screen "Point_1" 800x480, template "Main"
   TextField "Text field_1" at 0,2 size 547x23; Text 'Таблица настройки зависимостей дозы от мутность для линии 1'
   TextField "Text field_12" at 566,23 size 71x23; Text 'Запрос:'
   IOField "I/O field_4" at 653,22 size 66x25; FormatPattern 999.99
      ProcessValue <- "Ponts_1_DB_REQ"
   TextField "Text field_4" at 566,46 size 84x23; Text 'Команда:'
   IOField "I/O field_2" at 653,45 size 66x25; FormatPattern 999.99
      ProcessValue <- "Ponts_1_DB_Value"
   TextField "Text field_40" at 566,69 size 84x23; Text 'Датчик:'
   IOField "I/O field_24" at 653,68 size 66x25; FormatPattern 999.99
      ProcessValue <- "AIx_DB_Trans_1_Result"
   Rectangle "Rectangle_1" at 142,113 size 111x147
      Appearance <- "Ponts_1_DB_Now{1}"
   TextField "Text field_3" at 164,141 size 67x20; Text 'мутность'
   TextField "Text field_5" at 179,196 size 37x20; Text 'доза'
   TextField "Text field_11" at 142,115 size 95x25; Text 'Точка 1'
   Button "Button_1" at 223,113 size 30x30; TextOff 'Text'; Authorization "Operator"; PictureList "on_off_1"
      on Click: InvertBit("Ponts_1_DB_PLF_1_Use")
      ProcessValue <- "Ponts_1_DB_PLF_1_Use"
   IOField "I/O field_16" at 157,160 size 82x40; Authorization "Operator"; FormatPattern 999.99
      ProcessValue <- "Ponts_1_DB_PLF_1_High"
   IOField "I/O field_17" at 157,216 size 82x40; Authorization "Operator"; FormatPattern 999.99
      ProcessValue <- "Ponts_1_DB_PLF_1_Point_B"
   TextField "Text field_9" at 2,35 size 164x23; Text 'Минимальная доза'
   TextField "Text field_10" at 2,64 size 172x23; Text 'Максимальная доза'
   IOField "I/O field_1" at 181,33 size 70x30; Authorization "Operator"; FormatPattern 999.99
      ProcessValue <- "Ponts_1_DB_Min"
   IOField "I/O field_30" at 181,64 size 70x30; Authorization "Operator"; FormatPattern 999.99
      ProcessValue <- "Ponts_1_DB_Max"
   Rectangle "Rectangle_2" at 21,113 size 111x147
      Appearance <- "Ponts_1_DB_Now{0}"
   TextField "Text field_2" at 43,141 size 67x20; Text 'мутность'
   TextField "Text field_6" at 58,196 size 37x20; Text 'доза'
   TextField "Text field_7" at 21,115 size 95x25; Text 'Точка 0'
   Button "Button_2" at 102,113 size 30x30; TextOff 'Text'; Authorization "Operator"; PictureList "on_off_1"
      on Click: InvertBit("Ponts_1_DB_PLF_0_Use")
      ProcessValue <- "Ponts_1_DB_PLF_0_Use"
   IOField "I/O field_3" at 36,160 size 82x40; Authorization "Operator"; FormatPattern 999.99
      ProcessValue <- "Ponts_1_DB_PLF_0_High"
   IOField "I/O field_5" at 36,216 size 82x40; Authorization "Operator"; FormatPattern 999.99
      ProcessValue <- "Ponts_1_DB_PLF_0_Point_B"
   Rectangle "Rectangle_3" at 264,114 size 111x147
      Appearance <- "Ponts_1_DB_Now{2}"
   TextField "Text field_8" at 286,142 size 67x20; Text 'мутность'
   TextField "Text field_13" at 301,197 size 37x20; Text 'доза'
   TextField "Text field_14" at 264,116 size 95x25; Text 'Точка 2'
   Button "Button_3" at 345,114 size 30x30; TextOff 'Text'; Authorization "Operator"; PictureList "on_off_1"
      on Click: InvertBit("Ponts_1_DB_PLF_2_Use")
      ProcessValue <- "Ponts_1_DB_PLF_2_Use"
   IOField "I/O field_6" at 279,161 size 82x40; Authorization "Operator"; FormatPattern 999.99
      ProcessValue <- "Ponts_1_DB_PLF_2_High"
   IOField "I/O field_7" at 279,217 size 82x40; Authorization "Operator"; FormatPattern 999.99
      ProcessValue <- "Ponts_1_DB_PLF_2_Point_B"
   Rectangle "Rectangle_4" at 386,115 size 111x147
      Appearance <- "Ponts_1_DB_Now{3}"
   TextField "Text field_15" at 408,143 size 67x20; Text 'мутность'
   TextField "Text field_16" at 423,198 size 37x20; Text 'доза'
   TextField "Text field_17" at 386,117 size 95x25; Text 'Точка 3'
   Button "Button_4" at 467,115 size 30x30; TextOff 'Text'; Authorization "Operator"; PictureList "on_off_1"
      on Click: InvertBit("Ponts_1_DB_PLF_3_Use")
      ProcessValue <- "Ponts_1_DB_PLF_3_Use"
   IOField "I/O field_8" at 401,162 size 82x40; Authorization "Operator"; FormatPattern 999.99
      ProcessValue <- "Ponts_1_DB_PLF_3_High"
   IOField "I/O field_9" at 401,218 size 82x40; Authorization "Operator"; FormatPattern 999.99
      ProcessValue <- "Ponts_1_DB_PLF_3_Point_B"
   Rectangle "Rectangle_5" at 142,287 size 111x147
      Appearance <- "Ponts_1_DB_Now{5}"
   TextField "Text field_18" at 164,315 size 67x20; Text 'мутность'
   TextField "Text field_19" at 179,370 size 37x20; Text 'доза'
   TextField "Text field_20" at 142,289 size 95x25; Text 'Точка 5'
   Button "Button_5" at 223,287 size 30x30; TextOff 'Text'; Authorization "Operator"; PictureList "on_off_1"
      on Click: InvertBit("Ponts_1_DB_PLF_5_Use")
      ProcessValue <- "Ponts_1_DB_PLF_5_Use"
   IOField "I/O field_10" at 157,334 size 82x40; Authorization "Operator"; FormatPattern 999.99
      ProcessValue <- "Ponts_1_DB_PLF_5_High"
   IOField "I/O field_11" at 157,390 size 82x40; Authorization "Operator"; FormatPattern 999.99
      ProcessValue <- "Ponts_1_DB_PLF_5_Point_B"
   Rectangle "Rectangle_6" at 21,287 size 111x147
      Appearance <- "Ponts_1_DB_Now{4}"
   TextField "Text field_21" at 43,315 size 67x20; Text 'мутность'
   TextField "Text field_22" at 58,370 size 37x20; Text 'доза'
   TextField "Text field_23" at 21,289 size 95x25; Text 'Точка 4'
   Button "Button_6" at 102,287 size 30x30; TextOff 'Text'; Authorization "Operator"; PictureList "on_off_1"
      on Click: InvertBit("Ponts_1_DB_PLF_4_Use")
      ProcessValue <- "Ponts_1_DB_PLF_4_Use"
   IOField "I/O field_12" at 36,334 size 82x40; Authorization "Operator"; FormatPattern 999.99
      ProcessValue <- "Ponts_1_DB_PLF_4_High"
   IOField "I/O field_13" at 36,390 size 82x40; Authorization "Operator"; FormatPattern 999.99
      ProcessValue <- "Ponts_1_DB_PLF_4_Point_B"
   Rectangle "Rectangle_7" at 264,288 size 111x147
      Appearance <- "Ponts_1_DB_Now{6}"
   TextField "Text field_24" at 286,316 size 67x20; Text 'мутность'
   TextField "Text field_25" at 301,371 size 37x20; Text 'доза'
   TextField "Text field_26" at 264,290 size 95x25; Text 'Точка 6'
   Button "Button_7" at 345,288 size 30x30; TextOff 'Text'; Authorization "Operator"; PictureList "on_off_1"
      on Click: InvertBit("Ponts_1_DB_PLF_6_Use")
      ProcessValue <- "Ponts_1_DB_PLF_6_Use"
   IOField "I/O field_14" at 279,335 size 82x40; Authorization "Operator"; FormatPattern 999.99
      ProcessValue <- "Ponts_1_DB_PLF_6_High"
   IOField "I/O field_15" at 279,391 size 82x40; Authorization "Operator"; FormatPattern 999.99
      ProcessValue <- "Ponts_1_DB_PLF_6_Point_B"
   Rectangle "Rectangle_8" at 386,289 size 111x147
      Appearance <- "Ponts_1_DB_Now{7}"
   TextField "Text field_27" at 408,317 size 67x20; Text 'мутность'
   TextField "Text field_28" at 423,372 size 37x20; Text 'доза'
   TextField "Text field_29" at 386,291 size 95x25; Text 'Точка 7'
   Button "Button_8" at 467,289 size 30x30; TextOff 'Text'; Authorization "Operator"; PictureList "on_off_1"
      on Click: InvertBit("Ponts_1_DB_PLF_7_Use")
      ProcessValue <- "Ponts_1_DB_PLF_7_Use"
   IOField "I/O field_18" at 401,336 size 82x40; Authorization "Operator"; FormatPattern 999.99
      ProcessValue <- "Ponts_1_DB_PLF_7_High"
   IOField "I/O field_19" at 401,392 size 82x40; Authorization "Operator"; FormatPattern 999.99
      ProcessValue <- "Ponts_1_DB_PLF_7_Point_B"

screen "Point_2" 800x480, template "Main"
   TextField "Text field_1" at 0,2 size 547x23; Text 'Таблица настройки зависимостей дозы от мутность для линии 2'
   TextField "Text field_12" at 566,23 size 71x23; Text 'Запрос:'
   IOField "I/O field_4" at 653,22 size 66x25; FormatPattern 999.99
      ProcessValue <- "Ponts_2_DB_REQ"
   TextField "Text field_4" at 566,46 size 84x23; Text 'Команда:'
   IOField "I/O field_2" at 653,45 size 66x25; FormatPattern 999.99
      ProcessValue <- "Ponts_2_DB_Value"
   TextField "Text field_40" at 566,69 size 84x23; Text 'Датчик:'
   IOField "I/O field_24" at 653,68 size 66x25; FormatPattern 999.99
      ProcessValue <- "AIx_DB_Trans_2_Result"
   Rectangle "Rectangle_1" at 142,113 size 111x147
      Appearance <- "Ponts_2_DB_Now{1}"
   TextField "Text field_3" at 164,141 size 67x20; Text 'мутность'
   TextField "Text field_5" at 179,196 size 37x20; Text 'доза'
   TextField "Text field_11" at 142,115 size 95x25; Text 'Точка 1'
   Button "Button_1" at 223,113 size 30x30; TextOff 'Text'; Authorization "Operator"; PictureList "on_off_1"
      on Click: InvertBit("Ponts_2_DB_PLF_1_Use")
      ProcessValue <- "Ponts_2_DB_PLF_1_Use"
   IOField "I/O field_16" at 157,160 size 82x40; Authorization "Operator"; FormatPattern 999.99
      ProcessValue <- "Ponts_2_DB_PLF_1_High"
   IOField "I/O field_17" at 157,216 size 82x40; Authorization "Operator"; FormatPattern 999.99
      ProcessValue <- "Ponts_2_DB_PLF_1_Point_B"
   TextField "Text field_9" at 2,35 size 164x23; Text 'Минимальная доза'
   TextField "Text field_10" at 2,64 size 172x23; Text 'Максимальная доза'
   IOField "I/O field_1" at 181,33 size 70x30; Authorization "Operator"; FormatPattern 999.99
      ProcessValue <- "Ponts_2_DB_Min"
   IOField "I/O field_30" at 181,64 size 70x30; Authorization "Operator"; FormatPattern 999.99
      ProcessValue <- "Ponts_2_DB_Max"
   Rectangle "Rectangle_2" at 21,113 size 111x147
      Appearance <- "Ponts_2_DB_Now{0}"
   TextField "Text field_2" at 43,141 size 67x20; Text 'мутность'
   TextField "Text field_6" at 58,196 size 37x20; Text 'доза'
   TextField "Text field_7" at 21,115 size 95x25; Text 'Точка 0'
   Button "Button_2" at 102,113 size 30x30; TextOff 'Text'; Authorization "Operator"; PictureList "on_off_1"
      on Click: InvertBit("Ponts_2_DB_PLF_0_Use")
      ProcessValue <- "Ponts_2_DB_PLF_0_Use"
   IOField "I/O field_3" at 36,160 size 82x40; Authorization "Operator"; FormatPattern 999.99
      ProcessValue <- "Ponts_2_DB_PLF_0_High"
   IOField "I/O field_5" at 36,216 size 82x40; Authorization "Operator"; FormatPattern 999.99
      ProcessValue <- "Ponts_2_DB_PLF_0_Point_B"
   Rectangle "Rectangle_3" at 264,114 size 111x147
      Appearance <- "Ponts_2_DB_Now{2}"
   TextField "Text field_8" at 286,142 size 67x20; Text 'мутность'
   TextField "Text field_13" at 301,197 size 37x20; Text 'доза'
   TextField "Text field_14" at 264,116 size 95x25; Text 'Точка 2'
   Button "Button_3" at 345,114 size 30x30; TextOff 'Text'; Authorization "Operator"; PictureList "on_off_1"
      on Click: InvertBit("Ponts_2_DB_PLF_2_Use")
      ProcessValue <- "Ponts_2_DB_PLF_2_Use"
   IOField "I/O field_6" at 279,161 size 82x40; Authorization "Operator"; FormatPattern 999.99
      ProcessValue <- "Ponts_2_DB_PLF_2_High"
   IOField "I/O field_7" at 279,217 size 82x40; Authorization "Operator"; FormatPattern 999.99
      ProcessValue <- "Ponts_2_DB_PLF_2_Point_B"
   Rectangle "Rectangle_4" at 386,115 size 111x147
      Appearance <- "Ponts_2_DB_Now{3}"
   TextField "Text field_15" at 408,143 size 67x20; Text 'мутность'
   TextField "Text field_16" at 423,198 size 37x20; Text 'доза'
   TextField "Text field_17" at 386,117 size 95x25; Text 'Точка 3'
   Button "Button_4" at 467,115 size 30x30; TextOff 'Text'; Authorization "Operator"; PictureList "on_off_1"
      on Click: InvertBit("Ponts_2_DB_PLF_3_Use")
      ProcessValue <- "Ponts_2_DB_PLF_3_Use"
   IOField "I/O field_8" at 401,162 size 82x40; Authorization "Operator"; FormatPattern 999.99
      ProcessValue <- "Ponts_2_DB_PLF_3_High"
   IOField "I/O field_9" at 401,218 size 82x40; Authorization "Operator"; FormatPattern 999.99
      ProcessValue <- "Ponts_2_DB_PLF_3_Point_B"
   Rectangle "Rectangle_5" at 142,287 size 111x147
      Appearance <- "Ponts_2_DB_Now{5}"
   TextField "Text field_18" at 164,315 size 67x20; Text 'мутность'
   TextField "Text field_19" at 179,370 size 37x20; Text 'доза'
   TextField "Text field_20" at 142,289 size 95x25; Text 'Точка 5'
   Button "Button_5" at 223,287 size 30x30; TextOff 'Text'; Authorization "Operator"; PictureList "on_off_1"
      on Click: InvertBit("Ponts_2_DB_PLF_5_Use")
      ProcessValue <- "Ponts_2_DB_PLF_5_Use"
   IOField "I/O field_10" at 157,334 size 82x40; Authorization "Operator"; FormatPattern 999.99
      ProcessValue <- "Ponts_2_DB_PLF_5_High"
   IOField "I/O field_11" at 157,390 size 82x40; Authorization "Operator"; FormatPattern 999.99
      ProcessValue <- "Ponts_2_DB_PLF_5_Point_B"
   Rectangle "Rectangle_6" at 21,287 size 111x147
      Appearance <- "Ponts_2_DB_Now{4}"
   TextField "Text field_21" at 43,315 size 67x20; Text 'мутность'
   TextField "Text field_22" at 58,370 size 37x20; Text 'доза'
   TextField "Text field_23" at 21,289 size 95x25; Text 'Точка 4'
   Button "Button_6" at 102,287 size 30x30; TextOff 'Text'; Authorization "Operator"; PictureList "on_off_1"
      on Click: InvertBit("Ponts_2_DB_PLF_4_Use")
      ProcessValue <- "Ponts_2_DB_PLF_4_Use"
   IOField "I/O field_12" at 36,334 size 82x40; Authorization "Operator"; FormatPattern 999.99
      ProcessValue <- "Ponts_2_DB_PLF_4_High"
   IOField "I/O field_13" at 36,390 size 82x40; Authorization "Operator"; FormatPattern 999.99
      ProcessValue <- "Ponts_2_DB_PLF_4_Point_B"
   Rectangle "Rectangle_7" at 264,288 size 111x147
      Appearance <- "Ponts_2_DB_Now{6}"
   TextField "Text field_24" at 286,316 size 67x20; Text 'мутность'
   TextField "Text field_25" at 301,371 size 37x20; Text 'доза'
   TextField "Text field_26" at 264,290 size 95x25; Text 'Точка 6'
   Button "Button_7" at 345,288 size 30x30; TextOff 'Text'; Authorization "Operator"; PictureList "on_off_1"
      on Click: InvertBit("Ponts_2_DB_PLF_6_Use")
      ProcessValue <- "Ponts_2_DB_PLF_6_Use"
   IOField "I/O field_14" at 279,335 size 82x40; Authorization "Operator"; FormatPattern 999.99
      ProcessValue <- "Ponts_2_DB_PLF_6_High"
   IOField "I/O field_15" at 279,391 size 82x40; Authorization "Operator"; FormatPattern 999.99
      ProcessValue <- "Ponts_2_DB_PLF_6_Point_B"
   Rectangle "Rectangle_8" at 386,289 size 111x147
      Appearance <- "Ponts_2_DB_Now{7}"
   TextField "Text field_27" at 408,317 size 67x20; Text 'мутность'
   TextField "Text field_28" at 423,372 size 37x20; Text 'доза'
   TextField "Text field_29" at 386,291 size 95x25; Text 'Точка 7'
   Button "Button_8" at 467,289 size 30x30; TextOff 'Text'; Authorization "Operator"; PictureList "on_off_1"
      on Click: InvertBit("Ponts_2_DB_PLF_7_Use")
      ProcessValue <- "Ponts_2_DB_PLF_7_Use"
   IOField "I/O field_18" at 401,336 size 82x40; Authorization "Operator"; FormatPattern 999.99
      ProcessValue <- "Ponts_2_DB_PLF_7_High"
   IOField "I/O field_19" at 401,392 size 82x40; Authorization "Operator"; FormatPattern 999.99
      ProcessValue <- "Ponts_2_DB_PLF_7_Point_B"

screen "Mass_1" 800x480, template "Main"
   TextField "Text field_1" at 220,5 size 368x47; Text 'Статистика весов 1'
   Button "HmiScreenItemData_1" at 10,425 size 159x47; TextOn 'Система'; TextOff 'Прошлый месяц'; PictureOn "Navigates to System screens for KTP700 Basic+ PN 14.0.1.0"; PictureOff "Navigates to System screens for KTP700 Basic+ PN 14.0.1.0"
      on Release: ActivateScreen("Last_1", 0)
   Button "HmiScreenItemData_4" at 565,425 size 159x47; TextOn 'О нас'; TextOff 'Текущий месяц'; PictureOn "Navigates to System screens for KTP700 Basic+ PN 14.0.1.0"; PictureOff "Navigates to System screens for KTP700 Basic+ PN 14.0.1.0"
   IOField "I/O field_1" at 365,434 size 98x30; FormatPattern 99999.99
      ProcessValue <- "Statistics_DB_Today_1"
      Appearance <- "DIx_DB_Mass_1_Signal"
   TextField "Text field_17" at 257,435 size 93x27; Text 'Сегодня:'
   TextField "Text field_2" at 10,5 size 75x23; Text 'Сегодня'
   TextField "Text field_3" at 126,5 size 45x23; Text 'день'
   IOField "I/O field_2" at 88,3 size 37x30; FormatPattern 99
      ProcessValue <- "Statistics_DB_Today_Int"
      Appearance <- "DIx_DB_Mass_1_Signal"
   TextField "Text field_4" at 12,61 size 61x23; Text 'День 1'
   TextField "Text field_5" at 12,97 size 61x23; Text 'День 2'
   TextField "Text field_6" at 12,134 size 61x23; Text 'День 3'
   TextField "Text field_7" at 12,170 size 61x23; Text 'День 4'
   TextField "Text field_8" at 12,207 size 61x23; Text 'День 5'
   TextField "Text field_9" at 12,243 size 61x23; Text 'День 6'
   TextField "Text field_10" at 12,280 size 61x23; Text 'День 7'
   TextField "Text field_11" at 12,316 size 61x23; Text 'День 8'
   TextField "Text field_12" at 12,353 size 61x23; Text 'День 9'
   TextField "Text field_13" at 12,390 size 71x23; Text 'День 10'
   IOField "I/O field_8" at 90,59 size 80x27; Authorization "Operator"; FormatPattern 999999.9
      ProcessValue <- "Statistics_DB_Month_1{1}"
   IOField "I/O field_3" at 90,95 size 80x27; Authorization "Operator"; FormatPattern 999999.9
      ProcessValue <- "Statistics_DB_Month_1{2}"
   IOField "I/O field_4" at 90,132 size 80x27; Authorization "Operator"; FormatPattern 999999.9
      ProcessValue <- "Statistics_DB_Month_1{3}"
   IOField "I/O field_5" at 90,168 size 80x27; Authorization "Operator"; FormatPattern 999999.9
      ProcessValue <- "Statistics_DB_Month_1{4}"
   IOField "I/O field_6" at 90,205 size 80x27; Authorization "Operator"; FormatPattern 999999.9
      ProcessValue <- "Statistics_DB_Month_1{5}"
   IOField "I/O field_7" at 90,241 size 80x27; Authorization "Operator"; FormatPattern 999999.9
      ProcessValue <- "Statistics_DB_Month_1{6}"
   IOField "I/O field_9" at 90,278 size 80x27; Authorization "Operator"; FormatPattern 999999.9
      ProcessValue <- "Statistics_DB_Month_1{7}"
   IOField "I/O field_10" at 90,314 size 80x27; Authorization "Operator"; FormatPattern 999999.9
      ProcessValue <- "Statistics_DB_Month_1{8}"
   IOField "I/O field_11" at 90,351 size 80x27; Authorization "Operator"; FormatPattern 999999.9
      ProcessValue <- "Statistics_DB_Month_1{9}"
   IOField "I/O field_12" at 90,388 size 80x27; Authorization "Operator"; FormatPattern 999999.9
      ProcessValue <- "Statistics_DB_Month_1{10}"
   IOField "I/O field_13" at 565,316 size 159x30; FormatPattern 99999.9
      ProcessValue <- "Statistics_DB_Summ_1"
      Appearance <- "DIx_DB_Mass_1_Signal"
   TextField "Text field_14" at 595,284 size 100x27; Text 'За месяц:'
   TextField "Text field_15" at 611,359 size 67x27; Text 'Всего:'
   IOField "I/O field_14" at 565,387 size 159x30; FormatPattern 9999999.9
      ProcessValue <- "Statistics_DB_All_1"
      Appearance <- "DIx_DB_Mass_1_Signal"
   TextField "Text field_16" at 202,62 size 71x23; Text 'День 11'
   TextField "Text field_18" at 202,98 size 71x23; Text 'День 12'
   TextField "Text field_19" at 202,135 size 71x23; Text 'День 13'
   TextField "Text field_20" at 202,171 size 71x23; Text 'День 14'
   TextField "Text field_21" at 202,208 size 71x23; Text 'День 15'
   TextField "Text field_22" at 202,244 size 71x23; Text 'День 16'
   TextField "Text field_23" at 202,281 size 71x23; Text 'День 17'
   TextField "Text field_24" at 202,317 size 71x23; Text 'День 18'
   TextField "Text field_25" at 202,354 size 71x23; Text 'День 19'
   TextField "Text field_26" at 202,391 size 71x23; Text 'День 20'
   IOField "I/O field_15" at 280,60 size 80x27; Authorization "Operator"; FormatPattern 999999.9
      ProcessValue <- "Statistics_DB_Month_1{11}"
   IOField "I/O field_16" at 280,96 size 80x27; Authorization "Operator"; FormatPattern 999999.9
      ProcessValue <- "Statistics_DB_Month_1{12}"
   IOField "I/O field_17" at 280,133 size 80x27; Authorization "Operator"; FormatPattern 999999.9
      ProcessValue <- "Statistics_DB_Month_1{13}"
   IOField "I/O field_18" at 280,169 size 80x27; Authorization "Operator"; FormatPattern 999999.9
      ProcessValue <- "Statistics_DB_Month_1{14}"
   IOField "I/O field_19" at 280,206 size 80x27; Authorization "Operator"; FormatPattern 999999.9
      ProcessValue <- "Statistics_DB_Month_1{15}"
   IOField "I/O field_20" at 280,242 size 80x27; Authorization "Operator"; FormatPattern 999999.9
      ProcessValue <- "Statistics_DB_Month_1{16}"
   IOField "I/O field_21" at 280,279 size 80x27; Authorization "Operator"; FormatPattern 999999.9
      ProcessValue <- "Statistics_DB_Month_1{17}"
   IOField "I/O field_22" at 280,315 size 80x27; Authorization "Operator"; FormatPattern 999999.9
      ProcessValue <- "Statistics_DB_Month_1{18}"
   IOField "I/O field_23" at 280,352 size 80x27; Authorization "Operator"; FormatPattern 999999.9
      ProcessValue <- "Statistics_DB_Month_1{19}"
   IOField "I/O field_24" at 280,389 size 80x27; Authorization "Operator"; FormatPattern 999999.9
      ProcessValue <- "Statistics_DB_Month_1{20}"
   TextField "Text field_27" at 392,63 size 71x23; Text 'День 21'
   TextField "Text field_28" at 392,99 size 71x23; Text 'День 22'
   TextField "Text field_29" at 392,136 size 71x23; Text 'День 23'
   TextField "Text field_30" at 392,172 size 71x23; Text 'День 24'
   TextField "Text field_31" at 392,209 size 71x23; Text 'День 25'
   TextField "Text field_32" at 392,245 size 71x23; Text 'День 26'
   TextField "Text field_33" at 392,282 size 71x23; Text 'День 27'
   TextField "Text field_34" at 392,318 size 71x23; Text 'День 28'
   TextField "Text field_35" at 392,355 size 71x23; Text 'День 29'
   TextField "Text field_36" at 392,392 size 71x23; Text 'День 30'
   IOField "I/O field_25" at 470,61 size 80x27; Authorization "Operator"; FormatPattern 999999.9
      ProcessValue <- "Statistics_DB_Month_1{21}"
   IOField "I/O field_26" at 470,97 size 80x27; Authorization "Operator"; FormatPattern 999999.9
      ProcessValue <- "Statistics_DB_Month_1{22}"
   IOField "I/O field_27" at 470,134 size 80x27; Authorization "Operator"; FormatPattern 999999.9
      ProcessValue <- "Statistics_DB_Month_1{23}"
   IOField "I/O field_28" at 470,170 size 80x27; Authorization "Operator"; FormatPattern 999999.9
      ProcessValue <- "Statistics_DB_Month_1{24}"
   IOField "I/O field_29" at 470,207 size 80x27; Authorization "Operator"; FormatPattern 999999.9
      ProcessValue <- "Statistics_DB_Month_1{25}"
   IOField "I/O field_30" at 470,243 size 80x27; Authorization "Operator"; FormatPattern 999999.9
      ProcessValue <- "Statistics_DB_Month_1{26}"
   IOField "I/O field_31" at 470,280 size 80x27; Authorization "Operator"; FormatPattern 999999.9
      ProcessValue <- "Statistics_DB_Month_1{27}"
   IOField "I/O field_32" at 470,316 size 80x27; Authorization "Operator"; FormatPattern 999999.9
      ProcessValue <- "Statistics_DB_Month_1{28}"
   IOField "I/O field_33" at 470,353 size 80x27; Authorization "Operator"; FormatPattern 999999.9
      ProcessValue <- "Statistics_DB_Month_1{29}"
   IOField "I/O field_34" at 470,390 size 80x27; Authorization "Operator"; FormatPattern 999999.9
      ProcessValue <- "Statistics_DB_Month_1{30}"
   TextField "Text field_37" at 563,64 size 71x23; Text 'День 31'
   IOField "I/O field_35" at 644,62 size 80x27; Authorization "Operator"; FormatPattern 999999.9
      ProcessValue <- "Statistics_DB_Month_1{31}"

screen "Mass_2" 800x480, template "Main"
   TextField "Text field_1" at 220,5 size 368x47; Text 'Статистика весов 2'
   Button "HmiScreenItemData_1" at 10,425 size 159x47; TextOn 'Система'; TextOff 'Прошлый месяц'; PictureOn "Navigates to System screens for KTP700 Basic+ PN 14.0.1.0"; PictureOff "Navigates to System screens for KTP700 Basic+ PN 14.0.1.0"
      on Release: ActivateScreen("Last_2", 0)
   Button "HmiScreenItemData_4" at 565,425 size 159x47; TextOn 'О нас'; TextOff 'Текущий месяц'; PictureOn "Navigates to System screens for KTP700 Basic+ PN 14.0.1.0"; PictureOff "Navigates to System screens for KTP700 Basic+ PN 14.0.1.0"
   IOField "I/O field_1" at 365,434 size 98x30; FormatPattern 99999.99
      ProcessValue <- "Statistics_DB_Today_2"
      Appearance <- "DIx_DB_Mass_2_Signal"
   TextField "Text field_17" at 257,435 size 93x27; Text 'Сегодня:'
   TextField "Text field_3" at 10,5 size 75x23; Text 'Сегодня'
   TextField "Text field_4" at 126,5 size 45x23; Text 'день'
   IOField "I/O field_2" at 88,3 size 37x30; FormatPattern 99
      ProcessValue <- "Statistics_DB_Today_Int"
      Appearance <- "DIx_DB_Mass_1_Signal"
   TextField "Text field_5" at 12,61 size 61x23; Text 'День 1'
   TextField "Text field_6" at 12,97 size 61x23; Text 'День 2'
   TextField "Text field_7" at 12,134 size 61x23; Text 'День 3'
   TextField "Text field_8" at 12,170 size 61x23; Text 'День 4'
   TextField "Text field_9" at 12,207 size 61x23; Text 'День 5'
   TextField "Text field_10" at 12,243 size 61x23; Text 'День 6'
   TextField "Text field_11" at 12,280 size 61x23; Text 'День 7'
   TextField "Text field_12" at 12,316 size 61x23; Text 'День 8'
   TextField "Text field_13" at 12,353 size 61x23; Text 'День 9'
   TextField "Text field_14" at 12,390 size 71x23; Text 'День 10'
   IOField "I/O field_8" at 90,59 size 80x27; Authorization "Operator"; FormatPattern 999999.9
      ProcessValue <- "Statistics_DB_Month_2{1}"
   IOField "I/O field_3" at 90,95 size 80x27; Authorization "Operator"; FormatPattern 999999.9
      ProcessValue <- "Statistics_DB_Month_2{2}"
   IOField "I/O field_4" at 90,132 size 80x27; Authorization "Operator"; FormatPattern 999999.9
      ProcessValue <- "Statistics_DB_Month_2{3}"
   IOField "I/O field_5" at 90,168 size 80x27; Authorization "Operator"; FormatPattern 999999.9
      ProcessValue <- "Statistics_DB_Month_2{4}"
   IOField "I/O field_6" at 90,205 size 80x27; Authorization "Operator"; FormatPattern 999999.9
      ProcessValue <- "Statistics_DB_Month_2{5}"
   IOField "I/O field_7" at 90,241 size 80x27; Authorization "Operator"; FormatPattern 999999.9
      ProcessValue <- "Statistics_DB_Month_2{6}"
   IOField "I/O field_9" at 90,278 size 80x27; Authorization "Operator"; FormatPattern 999999.9
      ProcessValue <- "Statistics_DB_Month_2{7}"
   IOField "I/O field_10" at 90,314 size 80x27; Authorization "Operator"; FormatPattern 999999.9
      ProcessValue <- "Statistics_DB_Month_2{8}"
   IOField "I/O field_11" at 90,351 size 80x27; Authorization "Operator"; FormatPattern 999999.9
      ProcessValue <- "Statistics_DB_Month_2{9}"
   IOField "I/O field_12" at 90,388 size 80x27; Authorization "Operator"; FormatPattern 999999.9
      ProcessValue <- "Statistics_DB_Month_2{10}"
   IOField "I/O field_13" at 565,316 size 159x30; FormatPattern 99999.9
      ProcessValue <- "Statistics_DB_Summ_2"
      Appearance <- "DIx_DB_Mass_2_Signal"
   TextField "Text field_15" at 595,284 size 100x27; Text 'За месяц:'
   TextField "Text field_16" at 611,359 size 67x27; Text 'Всего:'
   IOField "I/O field_14" at 565,387 size 159x30; FormatPattern 9999999.9
      ProcessValue <- "Statistics_DB_All_2"
      Appearance <- "DIx_DB_Mass_2_Signal"
   TextField "Text field_18" at 202,62 size 71x23; Text 'День 11'
   TextField "Text field_19" at 202,98 size 71x23; Text 'День 12'
   TextField "Text field_20" at 202,135 size 71x23; Text 'День 13'
   TextField "Text field_21" at 202,171 size 71x23; Text 'День 14'
   TextField "Text field_22" at 202,208 size 71x23; Text 'День 15'
   TextField "Text field_23" at 202,244 size 71x23; Text 'День 16'
   TextField "Text field_24" at 202,281 size 71x23; Text 'День 17'
   TextField "Text field_25" at 202,317 size 71x23; Text 'День 18'
   TextField "Text field_26" at 202,354 size 71x23; Text 'День 19'
   TextField "Text field_27" at 202,391 size 71x23; Text 'День 20'
   IOField "I/O field_15" at 280,60 size 80x27; Authorization "Operator"; FormatPattern 999999.9
      ProcessValue <- "Statistics_DB_Month_2{11}"
   IOField "I/O field_16" at 280,96 size 80x27; Authorization "Operator"; FormatPattern 999999.9
      ProcessValue <- "Statistics_DB_Month_2{12}"
   IOField "I/O field_17" at 280,133 size 80x27; Authorization "Operator"; FormatPattern 999999.9
      ProcessValue <- "Statistics_DB_Month_2{13}"
   IOField "I/O field_18" at 280,169 size 80x27; Authorization "Operator"; FormatPattern 999999.9
      ProcessValue <- "Statistics_DB_Month_2{14}"
   IOField "I/O field_19" at 280,206 size 80x27; Authorization "Operator"; FormatPattern 999999.9
      ProcessValue <- "Statistics_DB_Month_2{15}"
   IOField "I/O field_20" at 280,242 size 80x27; Authorization "Operator"; FormatPattern 999999.9
      ProcessValue <- "Statistics_DB_Month_2{16}"
   IOField "I/O field_21" at 280,279 size 80x27; Authorization "Operator"; FormatPattern 999999.9
      ProcessValue <- "Statistics_DB_Month_2{17}"
   IOField "I/O field_22" at 280,315 size 80x27; Authorization "Operator"; FormatPattern 999999.9
      ProcessValue <- "Statistics_DB_Month_2{18}"
   IOField "I/O field_23" at 280,352 size 80x27; Authorization "Operator"; FormatPattern 999999.9
      ProcessValue <- "Statistics_DB_Month_2{19}"
   IOField "I/O field_24" at 280,389 size 80x27; Authorization "Operator"; FormatPattern 999999.9
      ProcessValue <- "Statistics_DB_Month_2{20}"
   TextField "Text field_28" at 392,63 size 71x23; Text 'День 21'
   TextField "Text field_29" at 392,99 size 71x23; Text 'День 22'
   TextField "Text field_30" at 392,136 size 71x23; Text 'День 23'
   TextField "Text field_31" at 392,172 size 71x23; Text 'День 24'
   TextField "Text field_32" at 392,209 size 71x23; Text 'День 25'
   TextField "Text field_33" at 392,245 size 71x23; Text 'День 26'
   TextField "Text field_34" at 392,282 size 71x23; Text 'День 27'
   TextField "Text field_35" at 392,318 size 71x23; Text 'День 28'
   TextField "Text field_36" at 392,355 size 71x23; Text 'День 29'
   TextField "Text field_37" at 392,392 size 71x23; Text 'День 30'
   IOField "I/O field_25" at 470,61 size 80x27; Authorization "Operator"; FormatPattern 999999.9
      ProcessValue <- "Statistics_DB_Month_2{21}"
   IOField "I/O field_26" at 470,97 size 80x27; Authorization "Operator"; FormatPattern 999999.9
      ProcessValue <- "Statistics_DB_Month_2{22}"
   IOField "I/O field_27" at 470,134 size 80x27; Authorization "Operator"; FormatPattern 999999.9
      ProcessValue <- "Statistics_DB_Month_2{23}"
   IOField "I/O field_28" at 470,170 size 80x27; Authorization "Operator"; FormatPattern 999999.9
      ProcessValue <- "Statistics_DB_Month_2{24}"
   IOField "I/O field_29" at 470,207 size 80x27; Authorization "Operator"; FormatPattern 999999.9
      ProcessValue <- "Statistics_DB_Month_2{25}"
   IOField "I/O field_30" at 470,243 size 80x27; Authorization "Operator"; FormatPattern 999999.9
      ProcessValue <- "Statistics_DB_Month_2{26}"
   IOField "I/O field_31" at 470,280 size 80x27; Authorization "Operator"; FormatPattern 999999.9
      ProcessValue <- "Statistics_DB_Month_2{27}"
   IOField "I/O field_32" at 470,316 size 80x27; Authorization "Operator"; FormatPattern 999999.9
      ProcessValue <- "Statistics_DB_Month_2{28}"
   IOField "I/O field_33" at 470,353 size 80x27; Authorization "Operator"; FormatPattern 999999.9
      ProcessValue <- "Statistics_DB_Month_2{29}"
   IOField "I/O field_34" at 470,390 size 80x27; Authorization "Operator"; FormatPattern 999999.9
      ProcessValue <- "Statistics_DB_Month_2{30}"
   TextField "Text field_38" at 563,64 size 71x23; Text 'День 31'
   IOField "I/O field_35" at 644,62 size 80x27; Authorization "Operator"; FormatPattern 999999.9
      ProcessValue <- "Statistics_DB_Month_2{31}"

screen "Last_1" 800x480, template "Main"
   TextField "Text field_1" at 220,5 size 368x47; Text 'Статистика весов 1'
   Button "HmiScreenItemData_1" at 10,425 size 159x47; TextOff 'Прошлый месяц'; TextOn 'Система'; Authorization "Admin"; PictureOff "Navigates to System screens for KTP700 Basic+ PN 14.0.1.0"; PictureOn "Navigates to System screens for KTP700 Basic+ PN 14.0.1.0"
   Button "HmiScreenItemData_4" at 565,425 size 159x47; TextOn 'О нас'; TextOff 'Текущий месяц'; PictureOn "Navigates to System screens for KTP700 Basic+ PN 14.0.1.0"; PictureOff "Navigates to System screens for KTP700 Basic+ PN 14.0.1.0"
      on Release: ActivateScreen("Mass_1", 0)
   TextField "Text field_4" at 12,61 size 61x23; Text 'День 1'
   TextField "Text field_5" at 12,97 size 61x23; Text 'День 2'
   TextField "Text field_6" at 12,134 size 61x23; Text 'День 3'
   TextField "Text field_7" at 12,170 size 61x23; Text 'День 4'
   TextField "Text field_8" at 12,207 size 61x23; Text 'День 5'
   TextField "Text field_9" at 12,243 size 61x23; Text 'День 6'
   TextField "Text field_10" at 12,280 size 61x23; Text 'День 7'
   TextField "Text field_11" at 12,316 size 61x23; Text 'День 8'
   TextField "Text field_12" at 12,353 size 61x23; Text 'День 9'
   TextField "Text field_13" at 12,390 size 71x23; Text 'День 10'
   IOField "I/O field_8" at 90,59 size 80x27; Authorization "Operator"; FormatPattern 999999.9
      ProcessValue <- "Statistics_DB_Last_M_1{1}"
   IOField "I/O field_3" at 90,95 size 80x27; Authorization "Operator"; FormatPattern 999999.9
      ProcessValue <- "Statistics_DB_Last_M_1{2}"
   IOField "I/O field_4" at 90,132 size 80x27; Authorization "Operator"; FormatPattern 999999.9
      ProcessValue <- "Statistics_DB_Last_M_1{3}"
   IOField "I/O field_5" at 90,168 size 80x27; Authorization "Operator"; FormatPattern 999999.9
      ProcessValue <- "Statistics_DB_Last_M_1{4}"
   IOField "I/O field_6" at 90,205 size 80x27; Authorization "Operator"; FormatPattern 999999.9
      ProcessValue <- "Statistics_DB_Last_M_1{5}"
   IOField "I/O field_7" at 90,241 size 80x27; Authorization "Operator"; FormatPattern 999999.9
      ProcessValue <- "Statistics_DB_Last_M_1{6}"
   IOField "I/O field_9" at 90,278 size 80x27; Authorization "Operator"; FormatPattern 999999.9
      ProcessValue <- "Statistics_DB_Last_M_1{7}"
   IOField "I/O field_10" at 90,314 size 80x27; Authorization "Operator"; FormatPattern 999999.9
      ProcessValue <- "Statistics_DB_Last_M_1{8}"
   IOField "I/O field_11" at 90,351 size 80x27; Authorization "Operator"; FormatPattern 999999.9
      ProcessValue <- "Statistics_DB_Last_M_1{9}"
   IOField "I/O field_12" at 90,388 size 80x27; Authorization "Operator"; FormatPattern 999999.9
      ProcessValue <- "Statistics_DB_Last_M_1{10}"
   IOField "I/O field_13" at 565,316 size 159x30; FormatPattern 99999.9
      ProcessValue <- "Statistics_DB_Last_Month_1"
      Appearance <- "DIx_DB_Mass_1_Signal"
   TextField "Text field_14" at 595,284 size 100x27; Text 'За месяц:'
   TextField "Text field_15" at 611,359 size 67x27; Text 'Всего:'
   IOField "I/O field_14" at 565,387 size 159x30; FormatPattern 9999999.9
      ProcessValue <- "Statistics_DB_All_1"
      Appearance <- "DIx_DB_Mass_1_Signal"
   TextField "Text field_16" at 202,62 size 71x23; Text 'День 11'
   TextField "Text field_18" at 202,98 size 71x23; Text 'День 12'
   TextField "Text field_19" at 202,135 size 71x23; Text 'День 13'
   TextField "Text field_20" at 202,171 size 71x23; Text 'День 14'
   TextField "Text field_21" at 202,208 size 71x23; Text 'День 15'
   TextField "Text field_22" at 202,244 size 71x23; Text 'День 16'
   TextField "Text field_23" at 202,281 size 71x23; Text 'День 17'
   TextField "Text field_24" at 202,317 size 71x23; Text 'День 18'
   TextField "Text field_25" at 202,354 size 71x23; Text 'День 19'
   TextField "Text field_26" at 202,391 size 71x23; Text 'День 20'
   IOField "I/O field_15" at 280,60 size 80x27; Authorization "Operator"; FormatPattern 999999.9
      ProcessValue <- "Statistics_DB_Last_M_1{11}"
   IOField "I/O field_16" at 280,96 size 80x27; Authorization "Operator"; FormatPattern 999999.9
      ProcessValue <- "Statistics_DB_Last_M_1{12}"
   IOField "I/O field_17" at 280,133 size 80x27; Authorization "Operator"; FormatPattern 999999.9
      ProcessValue <- "Statistics_DB_Last_M_1{13}"
   IOField "I/O field_18" at 280,169 size 80x27; Authorization "Operator"; FormatPattern 999999.9
      ProcessValue <- "Statistics_DB_Last_M_1{14}"
   IOField "I/O field_19" at 280,206 size 80x27; Authorization "Operator"; FormatPattern 999999.9
      ProcessValue <- "Statistics_DB_Last_M_1{15}"
   IOField "I/O field_20" at 280,242 size 80x27; Authorization "Operator"; FormatPattern 999999.9
      ProcessValue <- "Statistics_DB_Last_M_1{16}"
   IOField "I/O field_21" at 280,279 size 80x27; Authorization "Operator"; FormatPattern 999999.9
      ProcessValue <- "Statistics_DB_Last_M_1{17}"
   IOField "I/O field_22" at 280,315 size 80x27; Authorization "Operator"; FormatPattern 999999.9
      ProcessValue <- "Statistics_DB_Last_M_1{18}"
   IOField "I/O field_23" at 280,352 size 80x27; Authorization "Operator"; FormatPattern 999999.9
      ProcessValue <- "Statistics_DB_Last_M_1{19}"
   IOField "I/O field_24" at 280,389 size 80x27; Authorization "Operator"; FormatPattern 999999.9
      ProcessValue <- "Statistics_DB_Last_M_1{20}"
   TextField "Text field_27" at 392,63 size 71x23; Text 'День 21'
   TextField "Text field_28" at 392,99 size 71x23; Text 'День 22'
   TextField "Text field_29" at 392,136 size 71x23; Text 'День 23'
   TextField "Text field_30" at 392,172 size 71x23; Text 'День 24'
   TextField "Text field_31" at 392,209 size 71x23; Text 'День 25'
   TextField "Text field_32" at 392,245 size 71x23; Text 'День 26'
   TextField "Text field_33" at 392,282 size 71x23; Text 'День 27'
   TextField "Text field_34" at 392,318 size 71x23; Text 'День 28'
   TextField "Text field_35" at 392,355 size 71x23; Text 'День 29'
   TextField "Text field_36" at 392,392 size 71x23; Text 'День 30'
   IOField "I/O field_25" at 470,61 size 80x27; Authorization "Operator"; FormatPattern 999999.9
      ProcessValue <- "Statistics_DB_Last_M_1{21}"
   IOField "I/O field_26" at 470,97 size 80x27; Authorization "Operator"; FormatPattern 999999.9
      ProcessValue <- "Statistics_DB_Last_M_1{22}"
   IOField "I/O field_27" at 470,134 size 80x27; Authorization "Operator"; FormatPattern 999999.9
      ProcessValue <- "Statistics_DB_Last_M_1{23}"
   IOField "I/O field_28" at 470,170 size 80x27; Authorization "Operator"; FormatPattern 999999.9
      ProcessValue <- "Statistics_DB_Last_M_1{24}"
   IOField "I/O field_29" at 470,207 size 80x27; Authorization "Operator"; FormatPattern 999999.9
      ProcessValue <- "Statistics_DB_Last_M_1{25}"
   IOField "I/O field_30" at 470,243 size 80x27; Authorization "Operator"; FormatPattern 999999.9
      ProcessValue <- "Statistics_DB_Last_M_1{26}"
   IOField "I/O field_31" at 470,280 size 80x27; Authorization "Operator"; FormatPattern 999999.9
      ProcessValue <- "Statistics_DB_Last_M_1{27}"
   IOField "I/O field_32" at 470,316 size 80x27; Authorization "Operator"; FormatPattern 999999.9
      ProcessValue <- "Statistics_DB_Last_M_1{28}"
   IOField "I/O field_33" at 470,353 size 80x27; Authorization "Operator"; FormatPattern 999999.9
      ProcessValue <- "Statistics_DB_Last_M_1{29}"
   IOField "I/O field_34" at 470,390 size 80x27; Authorization "Operator"; FormatPattern 999999.9
      ProcessValue <- "Statistics_DB_Last_M_1{30}"
   TextField "Text field_37" at 563,64 size 71x23; Text 'День 31'
   IOField "I/O field_35" at 644,62 size 80x27; Authorization "Operator"; FormatPattern 999999.9
      ProcessValue <- "Statistics_DB_Last_M_1{31}"

screen "Last_2" 800x480, template "Main"
   TextField "Text field_1" at 220,5 size 368x47; Text 'Статистика весов 2'
   Button "HmiScreenItemData_1" at 10,425 size 159x47; TextOff 'Прошлый месяц'; TextOn 'Система'; PictureOn "Navigates to System screens for KTP700 Basic+ PN 14.0.1.0"; PictureOff "Navigates to System screens for KTP700 Basic+ PN 14.0.1.0"; Authorization "Admin"
   Button "HmiScreenItemData_4" at 565,425 size 159x47; TextOn 'О нас'; TextOff 'Текущий месяц'; PictureOn "Navigates to System screens for KTP700 Basic+ PN 14.0.1.0"; PictureOff "Navigates to System screens for KTP700 Basic+ PN 14.0.1.0"
      on Release: ActivateScreen("Mass_2", 0)
   TextField "Text field_5" at 12,61 size 61x23; Text 'День 1'
   TextField "Text field_6" at 12,97 size 61x23; Text 'День 2'
   TextField "Text field_7" at 12,134 size 61x23; Text 'День 3'
   TextField "Text field_8" at 12,170 size 61x23; Text 'День 4'
   TextField "Text field_9" at 12,207 size 61x23; Text 'День 5'
   TextField "Text field_10" at 12,243 size 61x23; Text 'День 6'
   TextField "Text field_11" at 12,280 size 61x23; Text 'День 7'
   TextField "Text field_12" at 12,316 size 61x23; Text 'День 8'
   TextField "Text field_13" at 12,353 size 61x23; Text 'День 9'
   TextField "Text field_14" at 12,390 size 71x23; Text 'День 10'
   IOField "I/O field_8" at 90,59 size 80x27; Authorization "Operator"; FormatPattern 999999.9
      ProcessValue <- "Statistics_DB_Last_M_2{1}"
   IOField "I/O field_3" at 90,95 size 80x27; Authorization "Operator"; FormatPattern 999999.9
      ProcessValue <- "Statistics_DB_Last_M_2{2}"
   IOField "I/O field_4" at 90,132 size 80x27; Authorization "Operator"; FormatPattern 999999.9
      ProcessValue <- "Statistics_DB_Last_M_2{3}"
   IOField "I/O field_5" at 90,168 size 80x27; Authorization "Operator"; FormatPattern 999999.9
      ProcessValue <- "Statistics_DB_Last_M_2{4}"
   IOField "I/O field_6" at 90,205 size 80x27; Authorization "Operator"; FormatPattern 999999.9
      ProcessValue <- "Statistics_DB_Last_M_2{5}"
   IOField "I/O field_7" at 90,241 size 80x27; Authorization "Operator"; FormatPattern 999999.9
      ProcessValue <- "Statistics_DB_Last_M_2{6}"
   IOField "I/O field_9" at 90,278 size 80x27; Authorization "Operator"; FormatPattern 999999.9
      ProcessValue <- "Statistics_DB_Last_M_2{7}"
   IOField "I/O field_10" at 90,314 size 80x27; Authorization "Operator"; FormatPattern 999999.9
      ProcessValue <- "Statistics_DB_Last_M_2{8}"
   IOField "I/O field_11" at 90,351 size 80x27; Authorization "Operator"; FormatPattern 999999.9
      ProcessValue <- "Statistics_DB_Last_M_2{9}"
   IOField "I/O field_12" at 90,388 size 80x27; Authorization "Operator"; FormatPattern 999999.9
      ProcessValue <- "Statistics_DB_Last_M_2{10}"
   IOField "I/O field_13" at 565,316 size 159x30; FormatPattern 99999.9
      ProcessValue <- "Statistics_DB_Last_Month_2"
      Appearance <- "DIx_DB_Mass_2_Signal"
   TextField "Text field_15" at 595,284 size 100x27; Text 'За месяц:'
   TextField "Text field_16" at 611,359 size 67x27; Text 'Всего:'
   IOField "I/O field_14" at 565,387 size 159x30; FormatPattern 9999999.9
      ProcessValue <- "Statistics_DB_All_2"
      Appearance <- "DIx_DB_Mass_2_Signal"
   TextField "Text field_18" at 202,62 size 71x23; Text 'День 11'
   TextField "Text field_19" at 202,98 size 71x23; Text 'День 12'
   TextField "Text field_20" at 202,135 size 71x23; Text 'День 13'
   TextField "Text field_21" at 202,171 size 71x23; Text 'День 14'
   TextField "Text field_22" at 202,208 size 71x23; Text 'День 15'
   TextField "Text field_23" at 202,244 size 71x23; Text 'День 16'
   TextField "Text field_24" at 202,281 size 71x23; Text 'День 17'
   TextField "Text field_25" at 202,317 size 71x23; Text 'День 18'
   TextField "Text field_26" at 202,354 size 71x23; Text 'День 19'
   TextField "Text field_27" at 202,391 size 71x23; Text 'День 20'
   IOField "I/O field_15" at 280,60 size 80x27; Authorization "Operator"; FormatPattern 999999.9
      ProcessValue <- "Statistics_DB_Last_M_2{11}"
   IOField "I/O field_16" at 280,96 size 80x27; Authorization "Operator"; FormatPattern 999999.9
      ProcessValue <- "Statistics_DB_Last_M_2{12}"
   IOField "I/O field_17" at 280,133 size 80x27; Authorization "Operator"; FormatPattern 999999.9
      ProcessValue <- "Statistics_DB_Last_M_2{13}"
   IOField "I/O field_18" at 280,169 size 80x27; Authorization "Operator"; FormatPattern 999999.9
      ProcessValue <- "Statistics_DB_Last_M_2{14}"
   IOField "I/O field_19" at 280,206 size 80x27; Authorization "Operator"; FormatPattern 999999.9
      ProcessValue <- "Statistics_DB_Last_M_2{15}"
   IOField "I/O field_20" at 280,242 size 80x27; Authorization "Operator"; FormatPattern 999999.9
      ProcessValue <- "Statistics_DB_Last_M_2{16}"
   IOField "I/O field_21" at 280,279 size 80x27; Authorization "Operator"; FormatPattern 999999.9
      ProcessValue <- "Statistics_DB_Last_M_2{17}"
   IOField "I/O field_22" at 280,315 size 80x27; Authorization "Operator"; FormatPattern 999999.9
      ProcessValue <- "Statistics_DB_Last_M_2{18}"
   IOField "I/O field_23" at 280,352 size 80x27; Authorization "Operator"; FormatPattern 999999.9
      ProcessValue <- "Statistics_DB_Last_M_2{19}"
   IOField "I/O field_24" at 280,389 size 80x27; Authorization "Operator"; FormatPattern 999999.9
      ProcessValue <- "Statistics_DB_Last_M_2{20}"
   TextField "Text field_28" at 392,63 size 71x23; Text 'День 21'
   TextField "Text field_29" at 392,99 size 71x23; Text 'День 22'
   TextField "Text field_30" at 392,136 size 71x23; Text 'День 23'
   TextField "Text field_31" at 392,172 size 71x23; Text 'День 24'
   TextField "Text field_32" at 392,209 size 71x23; Text 'День 25'
   TextField "Text field_33" at 392,245 size 71x23; Text 'День 26'
   TextField "Text field_34" at 392,282 size 71x23; Text 'День 27'
   TextField "Text field_35" at 392,318 size 71x23; Text 'День 28'
   TextField "Text field_36" at 392,355 size 71x23; Text 'День 29'
   TextField "Text field_37" at 392,392 size 71x23; Text 'День 30'
   IOField "I/O field_25" at 470,61 size 80x27; Authorization "Operator"; FormatPattern 999999.9
      ProcessValue <- "Statistics_DB_Last_M_2{21}"
   IOField "I/O field_26" at 470,97 size 80x27; Authorization "Operator"; FormatPattern 999999.9
      ProcessValue <- "Statistics_DB_Last_M_2{22}"
   IOField "I/O field_27" at 470,134 size 80x27; Authorization "Operator"; FormatPattern 999999.9
      ProcessValue <- "Statistics_DB_Last_M_2{23}"
   IOField "I/O field_28" at 470,170 size 80x27; Authorization "Operator"; FormatPattern 999999.9
      ProcessValue <- "Statistics_DB_Last_M_2{24}"
   IOField "I/O field_29" at 470,207 size 80x27; Authorization "Operator"; FormatPattern 999999.9
      ProcessValue <- "Statistics_DB_Last_M_2{25}"
   IOField "I/O field_30" at 470,243 size 80x27; Authorization "Operator"; FormatPattern 999999.9
      ProcessValue <- "Statistics_DB_Last_M_2{26}"
   IOField "I/O field_31" at 470,280 size 80x27; Authorization "Operator"; FormatPattern 999999.9
      ProcessValue <- "Statistics_DB_Last_M_2{27}"
   IOField "I/O field_32" at 470,316 size 80x27; Authorization "Operator"; FormatPattern 999999.9
      ProcessValue <- "Statistics_DB_Last_M_2{28}"
   IOField "I/O field_33" at 470,353 size 80x27; Authorization "Operator"; FormatPattern 999999.9
      ProcessValue <- "Statistics_DB_Last_M_2{29}"
   IOField "I/O field_34" at 470,390 size 80x27; Authorization "Operator"; FormatPattern 999999.9
      ProcessValue <- "Statistics_DB_Last_M_2{30}"
   TextField "Text field_38" at 563,64 size 71x23; Text 'День 31'
   IOField "I/O field_35" at 644,62 size 80x27; Authorization "Operator"; FormatPattern 999999.9
      ProcessValue <- "Statistics_DB_Last_M_2{31}"

Template "Main" 800x480
   Button "Button_1" at 735,5 size 60x60; TextOff 'Text'; PictureOff "home_2"
      on Click: ActivateScreen("Root screen", 0)
   Button "Button_2" at 735,72 size 60x60; TextOff 'Text'; PictureOff "sett"
      on Click: ActivateScreen("SP", 0)
   Button "Button_3" at 735,140 size 60x60; TextOff 'Text'; PictureOff "weight"
      on Click: ActivateScreen("Wieght", 0)
   Button "Button_4" at 735,207 size 60x60; TextOff 'Text'; PictureOff "sett_1"
      on Click: ActivateScreen("Monitor", 0)
   Button "Button_5" at 735,275 size 60x60; TextOff 'Text'; PictureOff "home_1"; PictureList "Alarm"
      on Click: ActivateScreen("Alarms", 0)
      ProcessValue <- "Any_Alm"
   Button "Button_6" at 735,342 size 60x60; TextOff 'Text'; PictureOff "back"
      on Click: function_efd93a16()
   Button "Button_7" at 735,410 size 60x60; TextOff 'Text'; PictureOff "reset"
      on Click: SetBit("Reset_All")
*)